       #tempPositionOfPostfix := #tempPositionOfPostfix + 1;
       #tempPositionOfPrePostfix := #tempPositionOfPrePostfix + 1;
       WHILE (#tempPrePostfix[#tempPositionOfPrePostfix + 1]) <= #LGCODE_MTH_PRSR_NUMBER_9 AND
         (#tempPrePostfix[#tempPositionOfPrePostfix + 1] >= #LGCODE_MTH_PRSR_NUMBER_0) AND
         (#tempPositionOfPrePostfix < #tempMaxPositionOfPrePostfix) DO
         #tempPostfixNotation[#tempPositionOfPostfix - 1] :=
         #tempPostfixNotation[#tempPositionOfPostfix - 1] + (#tempPrePostfix[#tempPositionOfPrePostfix + 1] - #LGCODE_MTH_PRSR_NUMBER_0)
         / #tempDenominatorDecimalNumbers;
         #tempPositionOfPrePostfix := #tempPositionOfPrePostfix + 1;
         #tempDenominatorDecimalNumbers := #tempDenominatorDecimalNumbers * 10;
       END_WHILE;
       #tempDenominatorDecimalNumbers := 10;
       //Falls negative Zahl
       IF #tempNextPostfixNumberIsNegative = TRUE THEN
         #tempPostfixNotation[#tempPositionOfPostfix - 1] := #tempPostfixNotation[#tempPositionOfPostfix - 1] * (-1);
         #tempNextPostfixNumberIsNegative := FALSE;
       END_IF;
       #tempPositionDecimalNumbers[#tempNumberOfDecimalNo] := #tempPositionOfPostfix - 1;
       #tempNumberOfDecimalNo := #tempNumberOfDecimalNo + 1;
     ELSIF
       //Zwei oder mehr Zahlen hintereinander erkennen und Zehner-, Hunderter-, Tausender- Stelle bilden
       (#tempPrePostfix[#tempPositionOfPrePostfix] <= #LGCODE_MTH_PRSR_NUMBER_9) AND
       (#tempPrePostfix[#tempPositionOfPrePostfix] >= #LGCODE_MTH_PRSR_NUMBER_0) AND
       (#tempPrePostfix[#tempPositionOfPrePostfix + 1] <= #LGCODE_MTH_PRSR_NUMBER_9) AND
       (#tempPrePostfix[#tempPositionOfPrePostfix + 1] >= #LGCODE_MTH_PRSR_NUMBER_0) AND
       (#tempPositionOfPrePostfix < #tempMaxPositionOfPrePostfix) AND
       (#tempPositionOfPrePostfix <> 0)
     THEN
       #tempPostfixNotation[#tempPositionOfPostfix] := (#tempPrePostfix[#tempPositionOfPrePostfix] - #LGCODE_MTH_PRSR_NUMBER_0);
       #tempPositionOfPostfix := #tempPositionOfPostfix + 1;
       WHILE (#tempPrePostfix[#tempPositionOfPrePostfix + 1] <= #LGCODE_MTH_PRSR_NUMBER_9) AND
         (#tempPrePostfix[#tempPositionOfPrePostfix + 1] >= #LGCODE_MTH_PRSR_NUMBER_0) AND
         (#tempPositionOfPrePostfix < #tempMaxPositionOfPrePostfix) DO
         #tempPostfixNotation[#tempPositionOfPostfix - 1] :=
         #tempPostfixNotation[#tempPositionOfPostfix - 1] * #LGCODE_MTH_PRSR_MULTIPLIER_FOR_MULTI_DIGIT_NO +
         (#tempPrePostfix[#tempPositionOfPrePostfix + 1] - #LGCODE_MTH_PRSR_NUMBER_0);
         #tempPositionOfPrePostfix := #tempPositionOfPrePostfix + 1;
       END_WHILE;
       #tempPositionMultiDigitNumbers[#tempNumberOfMultiDigitNo] := #tempPositionOfPostfix - 1;
       #tempNumberOfMultiDigitNo := #tempNumberOfMultiDigitNo + 1;
       //Falls mehrstellige Kommazahl
       IF #tempPrePostfix[#tempPositionOfPrePostfix + 1] = #LGCODE_MTH_PRSR_DECIMAL_POINT THEN
         #tempPositionOfPrePostfix := #tempPositionOfPrePostfix + 1;
         WHILE (#tempPrePostfix[#tempPositionOfPrePostfix + 1] <= #LGCODE_MTH_PRSR_NUMBER_9) AND
           (#tempPrePostfix[#tempPositionOfPrePostfix + 1] >= #LGCODE_MTH_PRSR_NUMBER_0) AND
           (#tempPositionOfPrePostfix < #tempMaxPositionOfPrePostfix) DO
           #tempPostfixNotation[#tempPositionOfPostfix - 1] := #tempPostfixNotation[#tempPositionOfPostfix - 1] +
           (#tempPrePostfix[#tempPositionOfPrePostfix + 1] - #LGCODE_MTH_PRSR_NUMBER_0) / #tempDenominatorDecimalNumbers;
           #tempPositionOfPrePostfix := #tempPositionOfPrePostfix + 1;
           #tempDenominatorDecimalNumbers := #tempDenominatorDecimalNumbers * 10;
         END_WHILE;
         #tempDenominatorDecimalNumbers := 10;
         #tempPositionDecimalNumbers[#tempNumberOfDecimalNo] := #tempPositionOfPostfix - 1;
         #tempNumberOfDecimalNo := #tempNumberOfDecimalNo + 1;
       END_IF;
       //Falls negative Zahl
       IF #tempNextPostfixNumberIsNegative = TRUE THEN
         #tempPostfixNotation[#tempPositionOfPostfix - 1] := #tempPostfixNotation[#tempPositionOfPostfix - 1] * (-1);
         #tempNextPostfixNumberIsNegative := FALSE;
       END_IF;
     ELSIF
       //Zahlen in Postfix-Notation schreiben
       (#tempPrePostfix[#tempPositionOfPrePostfix] <= #LGCODE_MTH_PRSR_NUMBER_9) AND (#tempPrePostfix[#tempPositionOfPrePostfix] >= #LGCODE_MTH_PRSR_NUMBER_0)
     THEN
       #tempPostfixNotation[#tempPositionOfPostfix] := (#tempPrePostfix[#tempPositionOfPrePostfix] - #LGCODE_MTH_PRSR_NUMBER_0);
       #tempPositionOfPostfix := #tempPositionOfPostfix + 1;
       //Falls negative Zahl
       IF #tempNextPostfixNumberIsNegative = TRUE THEN
         #tempPostfixNotation[#tempPositionOfPostfix - 1] := #tempPostfixNotation[#tempPositionOfPostfix - 1] * (-1);
         #tempNextPostfixNumberIsNegative := FALSE;
       END_IF;
     ELSIF
       //negative Zahlen erkennen
       ((#tempPrePostfix[#tempPositionOfPrePostfix] = #LGCODE_MTH_PRSR_MINUS) AND

       ((#tempPrePostfix[#tempPositionOfPrePostfix + 1] >= #LGCODE_MTH_PRSR_NUMBER_0) AND
       (#tempPrePostfix[#tempPositionOfPrePostfix + 1] <= #LGCODE_MTH_PRSR_NUMBER_9)) AND

       ((#tempPrePostfix[#tempPositionOfPrePostfix - 1] = #LGCODE_MTH_PRSR_MINUS) OR
       (#tempPrePostfix[#tempPositionOfPrePostfix - 1] = #LGCODE_MTH_PRSR_TIMES) OR
       (#tempPrePostfix[#tempPositionOfPrePostfix - 1] = #LGCODE_MTH_PRSR_PLUS) OR
       (#tempPrePostfix[#tempPositionOfPrePostfix - 1] = #LGCODE_MTH_PRSR_MINUS) OR
       (#tempPrePostfix[#tempPositionOfPrePostfix - 1] = #LGCODE_MTH_PRSR_DIVIDE) OR
       (#tempPrePostfix[#tempPositionOfPrePostfix - 1] = #LGCODE_MTH_PRSR_OPEN_BRACKET) OR
       (#tempPrePostfix[#tempPositionOfPrePostfix - 1] = #LGCODE_MTH_PRSR_LOGICAL_OR) OR
       (#tempPrePostfix[#tempPositionOfPrePostfix - 1] = #LGCODE_MTH_PRSR_LOGICAL_AND) OR
       (#tempPrePostfix[#tempPositionOfPrePostfix - 1] = #LGCODE_MTH_PRSR_LOGICAL_GREATER) OR
       (#tempPrePostfix[#tempPositionOfPrePostfix - 1] = #LGCODE_MTH_PRSR_LOGICAL_LESS) OR
       (#tempPrePostfix[#tempPositionOfPrePostfix - 1] = #LGCODE_MTH_PRSR_LOGICAL_EQUAL) OR
       (#tempPrePostfix[#tempPositionOfPrePostfix - 1] = #LGCODE_MTH_PRSR_LOGICAL_GREATER_EQUAL) OR
       (#tempPrePostfix[#tempPositionOfPrePostfix - 1] = #LGCODE_MTH_PRSR_LOGICAL_LESS_EQUAL) OR
       (#tempPrePostfix[#tempPositionOfPrePostfix - 1] = #LGCODE_MTH_PRSR_LOGICAL_NOT_EQUAL) OR
       (#tempPrePostfix[#tempPositionOfPrePostfix - 1] = #LGCODE_MTH_PRSR_LOGICAL_NOT) OR
       (#tempPrePostfix[#tempPositionOfPrePostfix - 1] = #LGCODE_MTH_PRSR_TO_THE_POWER_OF) OR
       (#tempPositionOfPrePostfix = 1)))
     THEN
       #tempNextPostfixNumberIsNegative := TRUE;
     ELSIF
       //negative Klammerausdrücke erkennen
       (#tempPrePostfix[#tempPositionOfPrePostfix] = #LGCODE_MTH_PRSR_MINUS) AND

       (#tempPrePostfix[#tempPositionOfPrePostfix + 1] = #LGCODE_MTH_PRSR_OPEN_BRACKET) AND

       ((#tempPrePostfix[#tempPositionOfPrePostfix - 1] = #LGCODE_MTH_PRSR_TIMES) OR
       (#tempPrePostfix[#tempPositionOfPrePostfix - 1] = #LGCODE_MTH_PRSR_PLUS) OR
       (#tempPrePostfix[#tempPositionOfPrePostfix - 1] = #LGCODE_MTH_PRSR_MINUS) OR
       (#tempPrePostfix[#tempPositionOfPrePostfix - 1] = #LGCODE_MTH_PRSR_DIVIDE) OR
       (#tempPrePostfix[#tempPositionOfPrePostfix - 1] = #LGCODE_MTH_PRSR_OPEN_BRACKET) OR
       (#tempPrePostfix[#tempPositionOfPrePostfix - 1] = #LGCODE_MTH_PRSR_CHAR_N) OR
       (#tempPrePostfix[#tempPositionOfPrePostfix - 1] = #LGCODE_MTH_PRSR_CHAR_S) OR
       (#tempPrePostfix[#tempPositionOfPrePostfix - 1] = #LGCODE_MTH_PRSR_CHAR_R) OR
       (#tempPrePostfix[#tempPositionOfPrePostfix - 1] = #LGCODE_MTH_PRSR_CHAR_T) OR
       (#tempPrePostfix[#tempPositionOfPrePostfix - 1] = #LGCODE_MTH_PRSR_LOGICAL_OR) OR
       (#tempPrePostfix[#tempPositionOfPrePostfix - 1] = #LGCODE_MTH_PRSR_LOGICAL_AND) OR
       (#tempPrePostfix[#tempPositionOfPrePostfix - 1] = #LGCODE_MTH_PRSR_LOGICAL_GREATER) OR
       (#tempPrePostfix[#tempPositionOfPrePostfix - 1] = #LGCODE_MTH_PRSR_LOGICAL_LESS) OR
       (#tempPrePostfix[#tempPositionOfPrePostfix - 1] = #LGCODE_MTH_PRSR_LOGICAL_EQUAL) OR
       (#tempPrePostfix[#tempPositionOfPrePostfix - 1] = #LGCODE_MTH_PRSR_LOGICAL_GREATER_EQUAL) OR
       (#tempPrePostfix[#tempPositionOfPrePostfix - 1] = #LGCODE_MTH_PRSR_LOGICAL_LESS_EQUAL) OR
       (#tempPrePostfix[#tempPositionOfPrePostfix - 1] = #LGCODE_MTH_PRSR_LOGICAL_NOT_EQUAL) OR
       (#tempPrePostfix[#tempPositionOfPrePostfix - 1] = #LGCODE_MTH_PRSR_LOGICAL_NOT) OR
       (#tempPrePostfix[#tempPositionOfPrePostfix - 1] = #LGCODE_MTH_PRSR_TO_THE_POWER_OF) OR
       (#tempPositionOfPrePostfix = 1))
     THEN
       #tempPositionOfNegBrackets[#tempNumberOfNegBrackets] := #tempPositionOfOperatorStack;
       #tempNumberOfNegBrackets := #tempNumberOfNegBrackets + 1;
     ELSIF
       //negative mathematische Funktion erkennen
       (#tempPrePostfix[#tempPositionOfPrePostfix] = #LGCODE_MTH_PRSR_MINUS) AND

       ((#tempPrePostfix[#tempPositionOfPrePostfix + 1] = #LGCODE_MTH_PRSR_CHAR_C) OR
       (#tempPrePostfix[#tempPositionOfPrePostfix + 1] = #LGCODE_MTH_PRSR_CHAR_S)) AND

       ((#tempPrePostfix[#tempPositionOfPrePostfix - 1] = #LGCODE_MTH_PRSR_TIMES) OR
       (#tempPrePostfix[#tempPositionOfPrePostfix - 1] = #LGCODE_MTH_PRSR_PLUS) OR
       (#tempPrePostfix[#tempPositionOfPrePostfix - 1] = #LGCODE_MTH_PRSR_MINUS) OR
       (#tempPrePostfix[#tempPositionOfPrePostfix - 1] = #LGCODE_MTH_PRSR_DIVIDE) OR
       (#tempPrePostfix[#tempPositionOfPrePostfix - 1] = #LGCODE_MTH_PRSR_OPEN_BRACKET) OR
       (#tempPrePostfix[#tempPositionOfPrePostfix - 1] = #LGCODE_MTH_PRSR_LOGICAL_OR) OR
       (#tempPrePostfix[#tempPositionOfPrePostfix - 1] = #LGCODE_MTH_PRSR_LOGICAL_AND) OR
       (#tempPrePostfix[#tempPositionOfPrePostfix - 1] = #LGCODE_MTH_PRSR_LOGICAL_GREATER) OR
       (#tempPrePostfix[#tempPositionOfPrePostfix - 1] = #LGCODE_MTH_PRSR_LOGICAL_LESS) OR
       (#tempPrePostfix[#tempPositionOfPrePostfix - 1] = #LGCODE_MTH_PRSR_LOGICAL_EQUAL) OR
       (#tempPrePostfix[#tempPositionOfPrePostfix - 1] = #LGCODE_MTH_PRSR_LOGICAL_GREATER_EQUAL) OR
       (#tempPrePostfix[#tempPositionOfPrePostfix - 1] = #LGCODE_MTH_PRSR_LOGICAL_LESS_EQUAL) OR
       (#tempPrePostfix[#tempPositionOfPrePostfix - 1] = #LGCODE_MTH_PRSR_LOGICAL_NOT_EQUAL) OR
       (#tempPrePostfix[#tempPositionOfPrePostfix - 1] = #LGCODE_MTH_PRSR_LOGICAL_NOT) OR
       (#tempPrePostfix[#tempPositionOfPrePostfix - 1] = #LGCODE_MTH_PRSR_TO_THE_POWER_OF) OR
       (#tempPositionOfPrePostfix = 1))
     THEN
       #tempPositionOfNegFunctions[#tempNumberOfNegFunctions] := #tempPositionOfOperatorStack;
       #tempNumberOfNegFunctions := #tempNumberOfNegFunctions + 1;
     ELSIF
       //Zeichen je nach Bedingungen in Zeichenspeicher oder in Postfix-Notation schreiben
       //Zeichenspeicher leer, Zeichen in Zeichenspeicher schreiben
       (((#tempPrePostfix[#tempPositionOfPrePostfix] = #LGCODE_MTH_PRSR_LOGICAL_OR) OR
       (#tempPrePostfix[#tempPositionOfPrePostfix] = #LGCODE_MTH_PRSR_LOGICAL_AND) OR
       (#tempPrePostfix[#tempPositionOfPrePostfix] = #LGCODE_MTH_PRSR_LOGICAL_GREATER) OR
       (#tempPrePostfix[#tempPositionOfPrePostfix] = #LGCODE_MTH_PRSR_LOGICAL_LESS) OR
       (#tempPrePostfix[#tempPositionOfPrePostfix] = #LGCODE_MTH_PRSR_LOGICAL_EQUAL) OR
       (#tempPrePostfix[#tempPositionOfPrePostfix] = #LGCODE_MTH_PRSR_LOGICAL_GREATER_EQUAL) OR
       (#tempPrePostfix[#tempPositionOfPrePostfix] = #LGCODE_MTH_PRSR_LOGICAL_LESS_EQUAL) OR
       (#tempPrePostfix[#tempPositionOfPrePostfix] = #LGCODE_MTH_PRSR_LOGICAL_NOT_EQUAL) OR
       (#tempPrePostfix[#tempPositionOfPrePostfix] = #LGCODE_MTH_PRSR_LOGICAL_NOT) OR
       (#tempPrePostfix[#tempPositionOfPrePostfix] = #LGCODE_MTH_PRSR_TIMES) OR
       (#tempPrePostfix[#tempPositionOfPrePostfix] = #LGCODE_MTH_PRSR_DIVIDE) OR
       (#tempPrePostfix[#tempPositionOfPrePostfix] = #LGCODE_MTH_PRSR_PLUS) OR
       (#tempPrePostfix[#tempPositionOfPrePostfix] = #LGCODE_MTH_PRSR_MINUS)) AND
       (#tempPositionOfOperatorStack = 1))
     THEN
       #tempStackForOperators[#tempPositionOfOperatorStack] := #tempPrePostfix[#tempPositionOfPrePostfix];
       #tempPositionOfOperatorStack := #tempPositionOfOperatorStack + 1;
     ELSIF
       //letztes Zeichen boolesch und nächstes mathematisch
       //Zeichen in Zeichenspeicher speichern
       ((#tempStackForOperators[#tempPositionOfOperatorStack - 1] = #LGCODE_MTH_PRSR_LOGICAL_GREATER) OR
       (#tempStackForOperators[#tempPositionOfOperatorStack - 1] = #LGCODE_MTH_PRSR_LOGICAL_LESS) OR
       (#tempStackForOperators[#tempPositionOfOperatorStack - 1] = #LGCODE_MTH_PRSR_LOGICAL_GREATER_EQUAL) OR
       (#tempStackForOperators[#tempPositionOfOperatorStack - 1] = #LGCODE_MTH_PRSR_LOGICAL_LESS_EQUAL) OR
       (#tempStackForOperators[#tempPositionOfOperatorStack - 1] = #LGCODE_MTH_PRSR_LOGICAL_EQUAL) OR
       (#tempStackForOperators[#tempPositionOfOperatorStack - 1] = #LGCODE_MTH_PRSR_LOGICAL_NOT_EQUAL) OR
       (#tempStackForOperators[#tempPositionOfOperatorStack - 1] = #LGCODE_MTH_PRSR_LOGICAL_AND) OR
       (#tempStackForOperators[#tempPositionOfOperatorStack - 1] = #LGCODE_MTH_PRSR_LOGICAL_OR))
       AND
       ((#tempPrePostfix[#tempPositionOfPrePostfix] = #LGCODE_MTH_PRSR_PLUS) OR
       (#tempPrePostfix[#tempPositionOfPrePostfix] = #LGCODE_MTH_PRSR_MINUS) OR
       (#tempPrePostfix[#tempPositionOfPrePostfix] = #LGCODE_MTH_PRSR_TIMES) OR
       (#tempPrePostfix[#tempPositionOfPrePostfix] = #LGCODE_MTH_PRSR_DIVIDE) OR
       (#tempPrePostfix[#tempPositionOfPrePostfix] = #LGCODE_MTH_PRSR_OPEN_BRACKET))
     THEN
       #tempStackForOperators[#tempPositionOfOperatorStack] := #tempPrePostfix[#tempPositionOfPrePostfix];
       #tempPositionOfOperatorStack := #tempPositionOfOperatorStack + 1;
     ELSIF
       //letztes Zeichen mathematisch und nächstes boolesch
       //dann alle mathematischen Zeichen erst aus Zeichenspeicher holen
       ((#tempStackForOperators[#tempPositionOfOperatorStack - 1] = #LGCODE_MTH_PRSR_TIMES) OR
       (#tempStackForOperators[#tempPositionOfOperatorStack - 1] = #LGCODE_MTH_PRSR_DIVIDE) OR
       (#tempStackForOperators[#tempPositionOfOperatorStack - 1] = #LGCODE_MTH_PRSR_MINUS) OR
       (#tempStackForOperators[#tempPositionOfOperatorStack - 1] = #LGCODE_MTH_PRSR_PLUS) OR
       (#tempStackForOperators[#tempPositionOfOperatorStack - 1] = #LGCODE_MTH_PRSR_SINUS) OR
       (#tempStackForOperators[#tempPositionOfOperatorStack - 1] = #LGCODE_MTH_PRSR_COSINUS) OR
       (#tempStackForOperators[#tempPositionOfOperatorStack - 1] = #LGCODE_MTH_PRSR_SQUARE) OR
       (#tempStackForOperators[#tempPositionOfOperatorStack - 1] = #LGCODE_MTH_PRSR_SQUAREROOT))
       AND
       ((#tempPrePostfix[#tempPositionOfPrePostfix] = #LGCODE_MTH_PRSR_LOGICAL_GREATER_EQUAL) OR
       (#tempPrePostfix[#tempPositionOfPrePostfix] = #LGCODE_MTH_PRSR_LOGICAL_LESS_EQUAL) OR
       (#tempPrePostfix[#tempPositionOfPrePostfix] = #LGCODE_MTH_PRSR_LOGICAL_EQUAL) OR
       (#tempPrePostfix[#tempPositionOfPrePostfix] = #LGCODE_MTH_PRSR_LOGICAL_NOT_EQUAL) OR
       (#tempPrePostfix[#tempPositionOfPrePostfix] = #LGCODE_MTH_PRSR_LOGICAL_GREATER) OR
       (#tempPrePostfix[#tempPositionOfPrePostfix] = #LGCODE_MTH_PRSR_LOGICAL_LESS) OR
       (#tempPrePostfix[#tempPositionOfPrePostfix] = #LGCODE_MTH_PRSR_LOGICAL_AND) OR
       (#tempPrePostfix[#tempPositionOfPrePostfix] = #LGCODE_MTH_PRSR_LOGICAL_OR))
     THEN
       #tempPostfixNotation[#tempPositionOfPostfix] := #tempStackForOperators[#tempPositionOfOperatorStack - 1];
       #tempPositionOfPostfix := #tempPositionOfPostfix + 1;
       #tempPositionOfOperatorStack := #tempPositionOfOperatorStack - 1;
       IF (#tempStackForOperators[#tempPositionOfOperatorStack - 1] = #LGCODE_MTH_PRSR_PLUS) OR
         (#tempStackForOperators[#tempPositionOfOperatorStack - 1] = #LGCODE_MTH_PRSR_MINUS) OR
         (#tempStackForOperators[#tempPositionOfOperatorStack - 1] = #LGCODE_MTH_PRSR_TIMES) OR
         (#tempStackForOperators[#tempPositionOfOperatorStack - 1] = #LGCODE_MTH_PRSR_DIVIDE)
       THEN
         #tempPostfixNotation[#tempPositionOfPostfix] := #tempStackForOperators[#tempPositionOfOperatorStack - 1];
         #tempPositionOfPostfix := #tempPositionOfPostfix + 1;
         #tempPositionOfOperatorStack := #tempPositionOfOperatorStack - 1;
       END_IF;
       #tempStackForOperators[#tempPositionOfOperatorStack] := #tempPrePostfix[#tempPositionOfPrePostfix];
       #tempPositionOfOperatorStack := #tempPositionOfOperatorStack + 1;
     ELSIF
       //letztes Zeichen >/ >= / <=/ =/<> oder < Nächstes & oder | dann Zeichen erst aus Zeichenspeicher holen
       ((#tempStackForOperators[#tempPositionOfOperatorStack - 1] = #LGCODE_MTH_PRSR_LOGICAL_GREATER) OR
       (#tempStackForOperators[#tempPositionOfOperatorStack - 1] = #LGCODE_MTH_PRSR_LOGICAL_LESS) OR
       (#tempStackForOperators[#tempPositionOfOperatorStack - 1] = #LGCODE_MTH_PRSR_LOGICAL_GREATER_EQUAL) OR
       (#tempStackForOperators[#tempPositionOfOperatorStack - 1] = #LGCODE_MTH_PRSR_LOGICAL_LESS_EQUAL) OR
       (#tempStackForOperators[#tempPositionOfOperatorStack - 1] = #LGCODE_MTH_PRSR_LOGICAL_EQUAL) OR
       (#tempStackForOperators[#tempPositionOfOperatorStack - 1] = #LGCODE_MTH_PRSR_LOGICAL_NOT_EQUAL))
       AND
       ((#tempPrePostfix[#tempPositionOfPrePostfix] = #LGCODE_MTH_PRSR_LOGICAL_AND) OR
       (#tempPrePostfix[#tempPositionOfPrePostfix] = #LGCODE_MTH_PRSR_LOGICAL_OR))
     THEN
       #tempPostfixNotation[#tempPositionOfPostfix] := #tempStackForOperators[#tempPositionOfOperatorStack - 1];
       #tempPositionOfPostfix := #tempPositionOfPostfix + 1;
       #tempPositionOfOperatorStack := #tempPositionOfOperatorStack - 1;
       IF    //Falls nächstes Zeichen im Zeichenspeicher noch ein AND oder AND
         ((#tempStackForOperators[#tempPositionOfOperatorStack - 1] = #LGCODE_MTH_PRSR_LOGICAL_AND) OR
         (#tempStackForOperators[#tempPositionOfOperatorStack - 1] = #LGCODE_MTH_PRSR_LOGICAL_OR))
       THEN
         #tempPostfixNotation[#tempPositionOfPostfix] := #tempStackForOperators[#tempPositionOfOperatorStack - 1];
         #tempPositionOfPostfix := #tempPositionOfPostfix + 1;
         #tempPositionOfOperatorStack := #tempPositionOfOperatorStack - 1;
       END_IF;
       #tempStackForOperators[#tempPositionOfOperatorStack] := #tempPrePostfix[#tempPositionOfPrePostfix];
       #tempPositionOfOperatorStack := #tempPositionOfOperatorStack + 1;
     ELSIF
       //letztes Zeichen >/ < / >=/<= /<> /=  oder <  und Nächstes ein >/ >= / <=/ <>/ = oder < dann erst Zeichen aus Zeichenspeicher holen
       //und dann erst kommendes Zeichen in Stack schreiben
       ((#tempStackForOperators[#tempPositionOfOperatorStack - 1] = #LGCODE_MTH_PRSR_LOGICAL_GREATER) OR
       (#tempStackForOperators[#tempPositionOfOperatorStack - 1] = #LGCODE_MTH_PRSR_LOGICAL_LESS) OR
       (#tempStackForOperators[#tempPositionOfOperatorStack - 1] = #LGCODE_MTH_PRSR_LOGICAL_GREATER_EQUAL) OR
       (#tempStackForOperators[#tempPositionOfOperatorStack - 1] = #LGCODE_MTH_PRSR_LOGICAL_LESS_EQUAL) OR
       (#tempStackForOperators[#tempPositionOfOperatorStack - 1] = #LGCODE_MTH_PRSR_LOGICAL_NOT_EQUAL) OR
       (#tempStackForOperators[#tempPositionOfOperatorStack - 1] = #LGCODE_MTH_PRSR_LOGICAL_EQUAL))
       AND
       ((#tempPrePostfix[#tempPositionOfPrePostfix] = #LGCODE_MTH_PRSR_LOGICAL_GREATER) OR
       (#tempPrePostfix[#tempPositionOfPrePostfix] = #LGCODE_MTH_PRSR_LOGICAL_LESS) OR
       (#tempPrePostfix[#tempPositionOfPrePostfix] = #LGCODE_MTH_PRSR_LOGICAL_GREATER_EQUAL) OR
       (#tempPrePostfix[#tempPositionOfPrePostfix] = #LGCODE_MTH_PRSR_LOGICAL_LESS_EQUAL) OR
       (#tempPrePostfix[#tempPositionOfPrePostfix] = #LGCODE_MTH_PRSR_LOGICAL_NOT_EQUAL) OR
       (#tempPrePostfix[#tempPositionOfPrePostfix] = #LGCODE_MTH_PRSR_LOGICAL_EQUAL))
     THEN
       #tempPostfixNotation[#tempPositionOfPostfix] := #tempStackForOperators[#tempPositionOfOperatorStack - 1];
       #tempPositionOfPostfix := #tempPositionOfPostfix + 1;
       #tempPositionOfOperatorStack := #tempPositionOfOperatorStack - 1;
       #tempStackForOperators[#tempPositionOfOperatorStack] := #tempPrePostfix[#tempPositionOfPrePostfix];
       #tempPositionOfOperatorStack := #tempPositionOfOperatorStack + 1;
     ELSIF
       //letztes Zeichen & oder | und Nächstes > /< />= / <= /<> /=   oder < dann Zeichen in Zeichenspeicher schreiben
       ((#tempStackForOperators[#tempPositionOfOperatorStack - 1] = #LGCODE_MTH_PRSR_LOGICAL_AND) OR
       (#tempStackForOperators[#tempPositionOfOperatorStack - 1] = #LGCODE_MTH_PRSR_LOGICAL_OR))
       AND
       ((#tempPrePostfix[#tempPositionOfPrePostfix] = #LGCODE_MTH_PRSR_LOGICAL_GREATER) OR
       (#tempPrePostfix[#tempPositionOfPrePostfix] = #LGCODE_MTH_PRSR_LOGICAL_LESS) OR
       (#tempPrePostfix[#tempPositionOfPrePostfix] = #LGCODE_MTH_PRSR_LOGICAL_GREATER_EQUAL) OR
       (#tempPrePostfix[#tempPositionOfPrePostfix] = #LGCODE_MTH_PRSR_LOGICAL_LESS_EQUAL) OR
       (#tempPrePostfix[#tempPositionOfPrePostfix] = #LGCODE_MTH_PRSR_LOGICAL_NOT_EQUAL) OR
       (#tempPrePostfix[#tempPositionOfPrePostfix] = #LGCODE_MTH_PRSR_LOGICAL_EQUAL))
     THEN
       #tempStackForOperators[#tempPositionOfOperatorStack] := #tempPrePostfix[#tempPositionOfPrePostfix];
       #tempPositionOfOperatorStack := #tempPositionOfOperatorStack + 1;
     ELSIF
       //letztes Zeichen  & oder | und Nächstes & oder | dann Zeichen erst aus Zeichenspeicher holen
       ((#tempStackForOperators[#tempPositionOfOperatorStack - 1] = #LGCODE_MTH_PRSR_LOGICAL_AND) OR
       (#tempStackForOperators[#tempPositionOfOperatorStack - 1] = #LGCODE_MTH_PRSR_LOGICAL_OR))
       AND
       ((#tempPrePostfix[#tempPositionOfPrePostfix] = #LGCODE_MTH_PRSR_LOGICAL_AND) OR
       (#tempPrePostfix[#tempPositionOfPrePostfix] = #LGCODE_MTH_PRSR_LOGICAL_OR))
     THEN
       #tempPostfixNotation[#tempPositionOfPostfix] := #tempStackForOperators[#tempPositionOfOperatorStack - 1];
       #tempPositionOfPostfix := #tempPositionOfPostfix + 1;
       #tempPositionOfOperatorStack := #tempPositionOfOperatorStack - 1;
       #tempStackForOperators[#tempPositionOfOperatorStack] := #tempPrePostfix[#tempPositionOfPrePostfix];
       #tempPositionOfOperatorStack := #tempPositionOfOperatorStack + 1;

     ELSIF
       //! immer in Zeichenspeicher schreiben
       (#tempPrePostfix[#tempPositionOfPrePostfix] = #LGCODE_MTH_PRSR_LOGICAL_NOT)
     THEN
       #tempStackForOperators[#tempPositionOfOperatorStack] := #tempPrePostfix[#tempPositionOfPrePostfix];
       #tempPositionOfOperatorStack := #tempPositionOfOperatorStack + 1;
     ELSIF
       //bei kommenden Zeichen, ! aus Zeichenspeicher holen
       (#tempStackForOperators[#tempPositionOfOperatorStack - 1] = #LGCODE_MTH_PRSR_LOGICAL_NOT)
       AND
       ((#tempPrePostfix[#tempPositionOfPrePostfix] = #LGCODE_MTH_PRSR_LOGICAL_GREATER) OR
       (#tempPrePostfix[#tempPositionOfPrePostfix] = #LGCODE_MTH_PRSR_LOGICAL_LESS) OR
       (#tempPrePostfix[#tempPositionOfPrePostfix] = #LGCODE_MTH_PRSR_LOGICAL_GREATER_EQUAL) OR
       (#tempPrePostfix[#tempPositionOfPrePostfix] = #LGCODE_MTH_PRSR_LOGICAL_LESS_EQUAL) OR
       (#tempPrePostfix[#tempPositionOfPrePostfix] = #LGCODE_MTH_PRSR_LOGICAL_NOT_EQUAL) OR
       (#tempPrePostfix[#tempPositionOfPrePostfix] = #LGCODE_MTH_PRSR_LOGICAL_EQUAL) OR
       (#tempPrePostfix[#tempPositionOfPrePostfix] = #LGCODE_MTH_PRSR_LOGICAL_AND) OR
       (#tempPrePostfix[#tempPositionOfPrePostfix] = #LGCODE_MTH_PRSR_LOGICAL_OR) OR
       (#tempPrePostfix[#tempPositionOfPrePostfix] = #LGCODE_MTH_PRSR_TO_THE_POWER_OF) OR
       (#tempPrePostfix[#tempPositionOfPrePostfix] = #LGCODE_MTH_PRSR_PLUS) OR
       (#tempPrePostfix[#tempPositionOfPrePostfix] = #LGCODE_MTH_PRSR_MINUS) OR
       (#tempPrePostfix[#tempPositionOfPrePostfix] = #LGCODE_MTH_PRSR_TIMES) OR
       (#tempPrePostfix[#tempPositionOfPrePostfix] = #LGCODE_MTH_PRSR_DIVIDE) OR
       (#tempPrePostfix[#tempPositionOfPrePostfix] = #LGCODE_MTH_PRSR_SINUS) OR
       (#tempPrePostfix[#tempPositionOfPrePostfix] = #LGCODE_MTH_PRSR_COSINUS) OR
       (#tempPrePostfix[#tempPositionOfPrePostfix] = #LGCODE_MTH_PRSR_SQUARE) OR
       (#tempPrePostfix[#tempPositionOfPrePostfix] = #LGCODE_MTH_PRSR_SQUAREROOT))
     THEN
       #tempPostfixNotation[#tempPositionOfPostfix] := #tempStackForOperators[#tempPositionOfOperatorStack - 1];
       #tempPositionOfPostfix := #tempPositionOfPostfix + 1;
       #tempPositionOfOperatorStack := #tempPositionOfOperatorStack - 1;
       //damit ausräumendes Zeichen im nächsten Durchgang korrekt verarbeitet wird
       #tempPositionOfPrePostfix := #tempPositionOfPrePostfix - 1;
     ELSIF
       //^ (Exponential-Operator) bei nächstem Zeichen aus Zeichenspeicher holen
       ((#tempStackForOperators[#tempPositionOfOperatorStack - 1] = #LGCODE_MTH_PRSR_TO_THE_POWER_OF)
       AND
       ((#tempPrePostfix[#tempPositionOfPrePostfix] = #LGCODE_MTH_PRSR_LOGICAL_GREATER) OR
       (#tempPrePostfix[#tempPositionOfPrePostfix] = #LGCODE_MTH_PRSR_LOGICAL_LESS) OR
       (#tempPrePostfix[#tempPositionOfPrePostfix] = #LGCODE_MTH_PRSR_LOGICAL_GREATER_EQUAL) OR
       (#tempPrePostfix[#tempPositionOfPrePostfix] = #LGCODE_MTH_PRSR_LOGICAL_LESS_EQUAL) OR
       (#tempPrePostfix[#tempPositionOfPrePostfix] = #LGCODE_MTH_PRSR_LOGICAL_NOT_EQUAL) OR
       (#tempPrePostfix[#tempPositionOfPrePostfix] = #LGCODE_MTH_PRSR_LOGICAL_EQUAL) OR
       (#tempPrePostfix[#tempPositionOfPrePostfix] = #LGCODE_MTH_PRSR_LOGICAL_AND) OR
       (#tempPrePostfix[#tempPositionOfPrePostfix] = #LGCODE_MTH_PRSR_LOGICAL_OR) OR
       (#tempPrePostfix[#tempPositionOfPrePostfix] = #LGCODE_MTH_PRSR_TO_THE_POWER_OF) OR
       (#tempPrePostfix[#tempPositionOfPrePostfix] = #LGCODE_MTH_PRSR_PLUS) OR
       (#tempPrePostfix[#tempPositionOfPrePostfix] = #LGCODE_MTH_PRSR_MINUS) OR
       (#tempPrePostfix[#tempPositionOfPrePostfix] = #LGCODE_MTH_PRSR_TIMES) OR
       (#tempPrePostfix[#tempPositionOfPrePostfix] = #LGCODE_MTH_PRSR_DIVIDE)))
     THEN
       #tempPostfixNotation[#tempPositionOfPostfix] := #tempStackForOperators[#tempPositionOfOperatorStack - 1];
       #tempPositionOfPostfix := #tempPositionOfPostfix + 1;
       #tempPositionOfOperatorStack := #tempPositionOfOperatorStack - 1;
       //damit ausräumendes Zeichen im nächsten Durchgang korrekt verarbeitet wird
       #tempPositionOfPrePostfix := #tempPositionOfPrePostfix - 1;
     ELSIF
       //^ (Exponential-Operator) in Zeichenspeicher schreiben,
       //außer oberstes Zeichen ist Funktion oder NOT, ist weiter oben realisiert
       (#tempPrePostfix[#tempPositionOfPrePostfix] = #LGCODE_MTH_PRSR_TO_THE_POWER_OF)
     THEN
       #tempStackForOperators[#tempPositionOfOperatorStack] := #tempPrePostfix[#tempPositionOfPrePostfix];
       #tempPositionOfOperatorStack := #tempPositionOfOperatorStack + 1;
     ELSIF
       //letztes Zeichen * oder / Nächstes + oder - dann erst Zeichen aus Zeichenspeicher holen
       ((#tempStackForOperators[#tempPositionOfOperatorStack - 1] = #LGCODE_MTH_PRSR_TIMES) OR
       (#tempStackForOperators[#tempPositionOfOperatorStack - 1] = #LGCODE_MTH_PRSR_DIVIDE)) AND
       ((#tempPrePostfix[#tempPositionOfPrePostfix] = #LGCODE_MTH_PRSR_PLUS) OR
       (#tempPrePostfix[#tempPositionOfPrePostfix] = #LGCODE_MTH_PRSR_MINUS))
     THEN
       #tempPostfixNotation[#tempPositionOfPostfix] := #tempStackForOperators[#tempPositionOfOperatorStack - 1];
       #tempPositionOfPostfix := #tempPositionOfPostfix + 1;
       #tempPositionOfOperatorStack := #tempPositionOfOperatorStack - 1;
       IF    //Falls nächstes Zeichen im Zeichenspeicher noch ein + oder -
         ((#tempStackForOperators[#tempPositionOfOperatorStack - 1] = #LGCODE_MTH_PRSR_PLUS) OR
         (#tempStackForOperators[#tempPositionOfOperatorStack - 1] = #LGCODE_MTH_PRSR_MINUS))
       THEN
         #tempPostfixNotation[#tempPositionOfPostfix] := #tempStackForOperators[#tempPositionOfOperatorStack - 1];
         #tempPositionOfPostfix := #tempPositionOfPostfix + 1;
         #tempPositionOfOperatorStack := #tempPositionOfOperatorStack - 1;
       END_IF;
       #tempStackForOperators[#tempPositionOfOperatorStack] := #tempPrePostfix[#tempPositionOfPrePostfix];
       #tempPositionOfOperatorStack := #tempPositionOfOperatorStack + 1;
     ELSIF
       //letztes Zeichen  * oder / Nächstes ein * oder / dann erst Zeichen aus Zeichenspeicher holen
       //und dann erst kommendes Zeichen in Stack schreiben
       ((#tempStackForOperators[#tempPositionOfOperatorStack - 1] = #LGCODE_MTH_PRSR_TIMES) OR
       (#tempStackForOperators[#tempPositionOfOperatorStack - 1] = #LGCODE_MTH_PRSR_DIVIDE)) AND
       ((#tempPrePostfix[#tempPositionOfPrePostfix] = #LGCODE_MTH_PRSR_TIMES) OR
       (#tempPrePostfix[#tempPositionOfPrePostfix] = #LGCODE_MTH_PRSR_DIVIDE))
     THEN
       #tempPostfixNotation[#tempPositionOfPostfix] := #tempStackForOperators[#tempPositionOfOperatorStack - 1];
       #tempPositionOfPostfix := #tempPositionOfPostfix + 1;
       #tempPositionOfOperatorStack := #tempPositionOfOperatorStack - 1;
       #tempStackForOperators[#tempPositionOfOperatorStack] := #tempPrePostfix[#tempPositionOfPrePostfix];
       #tempPositionOfOperatorStack := #tempPositionOfOperatorStack + 1;
     ELSIF
       //letztes Zeichen ein + oder - und Nächstes * oder / dann Zeichen in Zeichenspeicher schreiben
       ((#tempStackForOperators[#tempPositionOfOperatorStack - 1] = #LGCODE_MTH_PRSR_PLUS) OR
       (#tempStackForOperators[#tempPositionOfOperatorStack - 1] = #LGCODE_MTH_PRSR_MINUS)) AND
       ((#tempPrePostfix[#tempPositionOfPrePostfix] = #LGCODE_MTH_PRSR_TIMES) OR
       (#tempPrePostfix[#tempPositionOfPrePostfix] = #LGCODE_MTH_PRSR_DIVIDE))
     THEN
       #tempStackForOperators[#tempPositionOfOperatorStack] := #tempPrePostfix[#tempPositionOfPrePostfix];
       #tempPositionOfOperatorStack := #tempPositionOfOperatorStack + 1;
     ELSIF
       //letztes Zeichen  + oder - und Nächstes + oder - dann Zeichen erst aus Zeichenspeicher holen
       ((#tempStackForOperators[#tempPositionOfOperatorStack - 1] = #LGCODE_MTH_PRSR_PLUS) OR
       (#tempStackForOperators[#tempPositionOfOperatorStack - 1] = #LGCODE_MTH_PRSR_MINUS)) AND
       ((#tempPrePostfix[#tempPositionOfPrePostfix] = #LGCODE_MTH_PRSR_PLUS) OR
       (#tempPrePostfix[#tempPositionOfPrePostfix] = #LGCODE_MTH_PRSR_MINUS))
     THEN
       #tempPostfixNotation[#tempPositionOfPostfix] := #tempStackForOperators[#tempPositionOfOperatorStack - 1];
       #tempPositionOfPostfix := #tempPositionOfPostfix + 1;
       #tempPositionOfOperatorStack := #tempPositionOfOperatorStack - 1;
       #tempStackForOperators[#tempPositionOfOperatorStack] := #tempPrePostfix[#tempPositionOfPrePostfix];
       #tempPositionOfOperatorStack := #tempPositionOfOperatorStack + 1;
     ELSIF
       //kommende Öffnende Klammer ( immer in Zeichenspeicher speichern
       (#tempPrePostfix[#tempPositionOfPrePostfix] = #LGCODE_MTH_PRSR_OPEN_BRACKET)
     THEN
       #tempStackForOperators[#tempPositionOfOperatorStack] := #LGCODE_MTH_PRSR_OPEN_BRACKET;
       #tempPositionOfOperatorStack := #tempPositionOfOperatorStack + 1;
     ELSIF
       //letztes Zeichen eine öffnende Klammer (, dann kommendes Zeichen in Zeichenspeicher schreiben
       (#tempStackForOperators[#tempPositionOfOperatorStack - 1] = #LGCODE_MTH_PRSR_OPEN_BRACKET)
       AND
       ((#tempPrePostfix[#tempPositionOfPrePostfix] = #LGCODE_MTH_PRSR_LOGICAL_GREATER) OR
       (#tempPrePostfix[#tempPositionOfPrePostfix] = #LGCODE_MTH_PRSR_LOGICAL_LESS) OR
       (#tempPrePostfix[#tempPositionOfPrePostfix] = #LGCODE_MTH_PRSR_LOGICAL_GREATER_EQUAL) OR
       (#tempPrePostfix[#tempPositionOfPrePostfix] = #LGCODE_MTH_PRSR_LOGICAL_LESS_EQUAL) OR
       (#tempPrePostfix[#tempPositionOfPrePostfix] = #LGCODE_MTH_PRSR_LOGICAL_EQUAL) OR
       (#tempPrePostfix[#tempPositionOfPrePostfix] = #LGCODE_MTH_PRSR_LOGICAL_AND) OR
       (#tempPrePostfix[#tempPositionOfPrePostfix] = #LGCODE_MTH_PRSR_LOGICAL_OR) OR
       (#tempPrePostfix[#tempPositionOfPrePostfix] = #LGCODE_MTH_PRSR_PLUS) OR
       (#tempPrePostfix[#tempPositionOfPrePostfix] = #LGCODE_MTH_PRSR_MINUS) OR
       (#tempPrePostfix[#tempPositionOfPrePostfix] = #LGCODE_MTH_PRSR_TIMES) OR
       (#tempPrePostfix[#tempPositionOfPrePostfix] = #LGCODE_MTH_PRSR_DIVIDE))
     THEN
       #tempStackForOperators[#tempPositionOfOperatorStack] := #tempPrePostfix[#tempPositionOfPrePostfix];
       #tempPositionOfOperatorStack := #tempPositionOfOperatorStack + 1;
     ELSIF
       //nächstes Zeichen ist eine schließende Klammer
       //alle Zeichen aus Zeichenspeicher bis zur öffnenden Klammer in Postfix-Notation schreiben
       (#tempPrePostfix[#tempPositionOfPrePostfix] = #LGCODE_MTH_PRSR_CLOSE_BRACKET)
     THEN
       WHILE (#tempStackForOperators[#tempPositionOfOperatorStack - 1] <> #LGCODE_MTH_PRSR_OPEN_BRACKET) DO
         #tempPostfixNotation[#tempPositionOfPostfix] := #tempStackForOperators[#tempPositionOfOperatorStack - 1];
         #tempStackForOperators[#tempPositionOfOperatorStack - 1] := 0;
         #tempPositionOfOperatorStack := #tempPositionOfOperatorStack - 1;
         #tempPositionOfPostfix := #tempPositionOfPostfix + 1;
         //Falls eine negative mathematische Funktion kommt
         IF (#tempPositionOfNegFunctions[#tempNumberOfNegFunctions - 1] = #tempPositionOfOperatorStack) THEN
           #tempPositionOfNegTerm[#tempNumberOfNegTerm] := #tempPositionOfPostfix;
           #tempPositionOfPostfix := #tempPositionOfPostfix + 1;
           #tempNumberOfNegTerm := #tempNumberOfNegTerm + 1;
           #tempNumberOfNegFunctions := #tempNumberOfNegFunctions - 1;
         END_IF;
       END_WHILE;
       #tempPositionOfOperatorStack := #tempPositionOfOperatorStack - 1;
       #tempStackForOperators[#tempPositionOfOperatorStack] := 0;    //öffnende Klammer löschen
       //negative Klammerausdrücke
       IF (#tempPositionOfNegBrackets[#tempNumberOfNegBrackets - 1] = #tempPositionOfOperatorStack) THEN
         #tempPositionOfNegTerm[#tempNumberOfNegTerm] := #tempPositionOfPostfix;
         #tempPositionOfPostfix := #tempPositionOfPostfix + 1;
         #tempNumberOfNegTerm := #tempNumberOfNegTerm + 1;
         #tempNumberOfNegBrackets := #tempNumberOfNegBrackets - 1;
       END_IF;
     ELSIF    //sqr Quadrat
       (#tempPrePostfix[#tempPositionOfPrePostfix] = #LGCODE_MTH_PRSR_CHAR_S) AND
       (#tempPrePostfix[#tempPositionOfPrePostfix + 1] = #LGCODE_MTH_PRSR_CHAR_Q) AND
       (#tempPrePostfix[#tempPositionOfPrePostfix + 2] = #LGCODE_MTH_PRSR_CHAR_R) AND
       (#tempPrePostfix[#tempPositionOfPrePostfix + 3] <> #LGCODE_MTH_PRSR_CHAR_T)
     THEN
       #tempStackForOperators[#tempPositionOfOperatorStack] := #LGCODE_MTH_PRSR_SQUARE;
       #tempPositionOfOperatorStack := #tempPositionOfOperatorStack + 1;
       #tempPositionOfPrePostfix := #tempPositionOfPrePostfix + 2;
     ELSIF    //sqrt Quadratwurzel
       (#tempPrePostfix[#tempPositionOfPrePostfix] = #LGCODE_MTH_PRSR_CHAR_S) AND
       (#tempPrePostfix[#tempPositionOfPrePostfix + 1] = #LGCODE_MTH_PRSR_CHAR_Q) AND
       (#tempPrePostfix[#tempPositionOfPrePostfix + 2] = #LGCODE_MTH_PRSR_CHAR_R) AND
       (#tempPrePostfix[#tempPositionOfPrePostfix + 3] = #LGCODE_MTH_PRSR_CHAR_T)
     THEN
       #tempStackForOperators[#tempPositionOfOperatorStack] := #LGCODE_MTH_PRSR_SQUAREROOT;
       #tempPositionOfOperatorStack := #tempPositionOfOperatorStack + 1;
       #tempPositionOfPrePostfix := #tempPositionOfPrePostfix + 3;
     ELSIF    //sin Sinus
       (#tempPrePostfix[#tempPositionOfPrePostfix] = #LGCODE_MTH_PRSR_CHAR_S) AND
       (#tempPrePostfix[#tempPositionOfPrePostfix + 1] = #LGCODE_MTH_PRSR_CHAR_I) AND
       (#tempPrePostfix[#tempPositionOfPrePostfix + 2] = #LGCODE_MTH_PRSR_CHAR_N)
     THEN
       #tempStackForOperators[#tempPositionOfOperatorStack] := #LGCODE_MTH_PRSR_SINUS;
       #tempPositionOfOperatorStack := #tempPositionOfOperatorStack + 1;
       #tempPositionOfPrePostfix := #tempPositionOfPrePostfix + 2;
     ELSIF    //cos Cosinus
       (#tempPrePostfix[#tempPositionOfPrePostfix] = #LGCODE_MTH_PRSR_CHAR_C) AND
       (#tempPrePostfix[#tempPositionOfPrePostfix + 1] = #LGCODE_MTH_PRSR_CHAR_O) AND
       (#tempPrePostfix[#tempPositionOfPrePostfix + 2] = #LGCODE_MTH_PRSR_CHAR_S)
     THEN
       #tempStackForOperators[#tempPositionOfOperatorStack] := #LGCODE_MTH_PRSR_COSINUS;
       #tempPositionOfOperatorStack := #tempPositionOfOperatorStack + 1;
       #tempPositionOfPrePostfix := #tempPositionOfPrePostfix + 2;
     ELSIF
       //letztes Zeichen im Stack ist eine mathematische Funktion und Nächstes ein Rechen-Operator
       //Funktion wird auch bei logischen Operatoren (außer bei NOT) ausgelsen, oben realisiert
       ((#tempStackForOperators[#tempPositionOfOperatorStack - 1] = #LGCODE_MTH_PRSR_COSINUS) OR
       (#tempStackForOperators[#tempPositionOfOperatorStack - 1] = #LGCODE_MTH_PRSR_SINUS) OR
       (#tempStackForOperators[#tempPositionOfOperatorStack - 1] = #LGCODE_MTH_PRSR_SQUARE) OR
       (#tempStackForOperators[#tempPositionOfOperatorStack - 1] = #LGCODE_MTH_PRSR_SQUAREROOT)) AND
       ((#tempPrePostfix[#tempPositionOfPrePostfix] = #LGCODE_MTH_PRSR_TIMES) OR
       (#tempPrePostfix[#tempPositionOfPrePostfix] = #LGCODE_MTH_PRSR_MINUS) OR
       (#tempPrePostfix[#tempPositionOfPrePostfix] = #LGCODE_MTH_PRSR_PLUS) OR
       (#tempPrePostfix[#tempPositionOfPrePostfix] = #LGCODE_MTH_PRSR_DIVIDE))
     THEN
       #tempPostfixNotation[#tempPositionOfPostfix] := #tempStackForOperators[#tempPositionOfOperatorStack - 1];
       #tempPositionOfPostfix := #tempPositionOfPostfix + 1;
       #tempPositionOfOperatorStack := #tempPositionOfOperatorStack - 1;
       //Falls die mathematische Funktion negative ist
       IF (#tempPositionOfNegFunctions[#tempNumberOfNegFunctions - 1] = #tempPositionOfOperatorStack) THEN
         #tempPositionOfNegTerm[#tempNumberOfNegTerm] := #tempPositionOfPostfix;
         #tempPositionOfPostfix := #tempPositionOfPostfix + 1;
         #tempNumberOfNegTerm := #tempNumberOfNegTerm + 1;
         #tempNumberOfNegFunctions := #tempNumberOfNegFunctions - 1;
       END_IF;
       #tempPositionOfPrePostfix := #tempPositionOfPrePostfix - 1;
     ELSE
       ;
     END_IF;
     //Wenn PrePostfix-Array komplett eingelesen, Zeichenspeicher vollständig leeren
     IF (#tempPositionOfPrePostfix = #tempMaxPositionOfPrePostfix) THEN
       WHILE (#tempPositionOfOperatorStack > 1) DO
         #tempPostfixNotation[#tempPositionOfPostfix] := #tempStackForOperators[#tempPositionOfOperatorStack - 1];
         #tempStackForOperators[#tempPositionOfOperatorStack - 1] := 0;
         #tempPositionOfOperatorStack := #tempPositionOfOperatorStack - 1;
         #tempPositionOfPostfix := #tempPositionOfPostfix + 1;
         //Falls die mathematische Funktion negative ist
         IF (#tempPositionOfNegFunctions[#tempNumberOfNegFunctions - 1] = #tempPositionOfOperatorStack) THEN
           #tempPositionOfNegTerm[#tempNumberOfNegTerm] := #tempPositionOfPostfix;
           #tempPositionOfPostfix := #tempPositionOfPostfix + 1;
           #tempNumberOfNegTerm := #tempNumberOfNegTerm + 1;
           #tempNumberOfNegFunctions := #tempNumberOfNegFunctions - 1;
         END_IF;
       END_WHILE;
     END_IF;
     #tempPositionOfPrePostfix := #tempPositionOfPrePostfix + 1;
     #tempMaxOfPostfixPosition := #tempPositionOfPostfix;
   END_WHILE;
   #tempPositionOfPostfix := 1;
   #tempNumberOfMultiDigitNo := 1;
   #tempNumberOfNegTerm := 1;

   //Auswertung
   WHILE (#tempPositionOfPostfix <= #tempMaxOfPostfixPosition) DO
     IF (#tempPositionOfPostfix = #tempPositionOfNegTerm[#tempNumberOfNegTerm]) THEN
       //Vorzeichen des Ergebnisses des Klammerausdruckes negieren
       #tempStackOfIntermediateResults[#tempPositionOfIntermediateResult - 1] :=
       #tempStackOfIntermediateResults[#tempPositionOfIntermediateResult - 1] * (-1);
       #tempNumberOfNegTerm := #tempNumberOfNegTerm + 1;
       //Auswertung Zahlen Zeichen usw.
     ELSIF
       //um mehrstellige Zahlen nicht mit den ASCII Codierungen für Operatoren und Funktionen zu verwechseln
       (#tempPositionOfPostfix = #tempPositionMultiDigitNumbers[#tempNumberOfMultiDigitNo])
     THEN
       #tempStackOfIntermediateResults[#tempPositionOfIntermediateResult] := #tempPostfixNotation[#tempPositionOfPostfix];
       #tempPositionOfIntermediateResult := #tempPositionOfIntermediateResult + 1;
       #tempNumberOfMultiDigitNo := #tempNumberOfMultiDigitNo + 1;
     ELSIF
       //Falls Kommazahlen, negative Zahlen kommen, Abfrage kommendes Zeichen ungleich + - * /
       (#tempPostfixNotation[#tempPositionOfPostfix] <> #LGCODE_MTH_PRSR_LOGICAL_GREATER) AND
       (#tempPostfixNotation[#tempPositionOfPostfix] <> #LGCODE_MTH_PRSR_LOGICAL_LESS) AND
       (#tempPostfixNotation[#tempPositionOfPostfix] <> #LGCODE_MTH_PRSR_LOGICAL_GREATER_EQUAL) AND
       (#tempPostfixNotation[#tempPositionOfPostfix] <> #LGCODE_MTH_PRSR_LOGICAL_LESS_EQUAL) AND
       (#tempPostfixNotation[#tempPositionOfPostfix] <> #LGCODE_MTH_PRSR_LOGICAL_AND) AND
       (#tempPostfixNotation[#tempPositionOfPostfix] <> #LGCODE_MTH_PRSR_LOGICAL_OR) AND
       (#tempPostfixNotation[#tempPositionOfPostfix] <> #LGCODE_MTH_PRSR_LOGICAL_NOT) AND
       (#tempPostfixNotation[#tempPositionOfPostfix] <> #LGCODE_MTH_PRSR_LOGICAL_NOT_EQUAL) AND
       (#tempPostfixNotation[#tempPositionOfPostfix] <> #LGCODE_MTH_PRSR_LOGICAL_EQUAL) AND
       (#tempPostfixNotation[#tempPositionOfPostfix] <> #LGCODE_MTH_PRSR_MINUS) AND
       (#tempPostfixNotation[#tempPositionOfPostfix] <> #LGCODE_MTH_PRSR_PLUS) AND
       (#tempPostfixNotation[#tempPositionOfPostfix] <> #LGCODE_MTH_PRSR_TIMES) AND
       (#tempPostfixNotation[#tempPositionOfPostfix] <> #LGCODE_MTH_PRSR_DIVIDE) AND
       (#tempPostfixNotation[#tempPositionOfPostfix] <> #LGCODE_MTH_PRSR_SQUARE) AND
       (#tempPostfixNotation[#tempPositionOfPostfix] <> #LGCODE_MTH_PRSR_SQUAREROOT) AND
       (#tempPostfixNotation[#tempPositionOfPostfix] <> #LGCODE_MTH_PRSR_SINUS) AND
       (#tempPostfixNotation[#tempPositionOfPostfix] <> #LGCODE_MTH_PRSR_COSINUS) AND
       (#tempPostfixNotation[#tempPositionOfPostfix] <> #LGCODE_MTH_PRSR_TO_THE_POWER_OF)
     THEN
       #tempStackOfIntermediateResults[#tempPositionOfIntermediateResult] :=
       #tempPostfixNotation[#tempPositionOfPostfix];
       #tempPositionOfIntermediateResult := #tempPositionOfIntermediateResult + 1;

       //Auswertung ob +, -, * oder / und eigentliche Berechnung des mathematischen Ausdrucks
     ELSIF (#tempPostfixNotation[#tempPositionOfPostfix] = #LGCODE_MTH_PRSR_PLUS) THEN
       #tempStackOfIntermediateResults[#tempPositionOfIntermediateResult - 2] :=
       #tempStackOfIntermediateResults[#tempPositionOfIntermediateResult - 2] +
       #tempStackOfIntermediateResults[#tempPositionOfIntermediateResult - 1];
       #tempPositionOfIntermediateResult := #tempPositionOfIntermediateResult - 1;
     ELSIF (#tempPostfixNotation[#tempPositionOfPostfix] = #LGCODE_MTH_PRSR_MINUS) THEN
       #tempStackOfIntermediateResults[#tempPositionOfIntermediateResult - 2] :=
       #tempStackOfIntermediateResults[#tempPositionOfIntermediateResult - 2] -
       #tempStackOfIntermediateResults[#tempPositionOfIntermediateResult - 1];
       #tempPositionOfIntermediateResult := #tempPositionOfIntermediateResult - 1;
     ELSIF (#tempPostfixNotation[#tempPositionOfPostfix] = #LGCODE_MTH_PRSR_TIMES) THEN
       #tempStackOfIntermediateResults[#tempPositionOfIntermediateResult - 2] :=
       #tempStackOfIntermediateResults[#tempPositionOfIntermediateResult - 2] *
       #tempStackOfIntermediateResults[#tempPositionOfIntermediateResult - 1];
       #tempPositionOfIntermediateResult := #tempPositionOfIntermediateResult - 1;
     ELSIF (#tempPostfixNotation[#tempPositionOfPostfix] = #LGCODE_MTH_PRSR_DIVIDE) THEN

       // Prüfen auf Division durch Null
       IF (#tempStackOfIntermediateResults[#tempPositionOfIntermediateResult - 1] <> 0.0) THEN
         #tempStackOfIntermediateResults[#tempPositionOfIntermediateResult - 2] :=
         #tempStackOfIntermediateResults[#tempPositionOfIntermediateResult - 2] /
         #tempStackOfIntermediateResults[#tempPositionOfIntermediateResult - 1];
       ELSE
         #LKinLang_CalcMathAndBool.errorID := #LGCODE_MTH_PRSR_ERR_ID_DIVISION_BY_ZERO;
         #LKinLang_CalcMathAndBool.finalResult := 0;

         RETURN;
       END_IF;

       #tempPositionOfIntermediateResult := #tempPositionOfIntermediateResult - 1;
       //Auswertung sqr
     ELSIF (#tempPostfixNotation[#tempPositionOfPostfix] = #LGCODE_MTH_PRSR_SQUARE) THEN
       #tempStackOfIntermediateResults[#tempPositionOfIntermediateResult - 1] :=
       #tempStackOfIntermediateResults[#tempPositionOfIntermediateResult - 1] ** 2;
       //Auswertung sqrt
     ELSIF (#tempPostfixNotation[#tempPositionOfPostfix] = #LGCODE_MTH_PRSR_SQUAREROOT) THEN

       // Prüfen auf negative Wurzel
       IF (#tempStackOfIntermediateResults[#tempPositionOfIntermediateResult - 1] < 0.0) THEN
         #LKinLang_CalcMathAndBool.errorID := #LGCODE_MTH_PRSR_ERR_ID_NEAGTIVE_SQUARE_ROOT_ARGUMENT;
         #LKinLang_CalcMathAndBool.finalResult := 0;

         RETURN;
       ELSE
         #tempStackOfIntermediateResults[#tempPositionOfIntermediateResult - 1] :=
         SQRT(IN := #tempStackOfIntermediateResults[#tempPositionOfIntermediateResult - 1]);
       END_IF;

       //Auswertung sin
     ELSIF (#tempPostfixNotation[#tempPositionOfPostfix] = #LGCODE_MTH_PRSR_SINUS) THEN
       #tempStackOfIntermediateResults[#tempPositionOfIntermediateResult - 1] :=
       SIN(IN := #tempStackOfIntermediateResults[#tempPositionOfIntermediateResult - 1] * #LGCODE_MTH_PRSR_PI / 180);
       //Auswertung cos
     ELSIF (#tempPostfixNotation[#tempPositionOfPostfix] = #LGCODE_MTH_PRSR_COSINUS) THEN
       #tempStackOfIntermediateResults[#tempPositionOfIntermediateResult - 1] :=
       COS(IN := #tempStackOfIntermediateResults[#tempPositionOfIntermediateResult - 1] * #LGCODE_MTH_PRSR_PI / 180);
       //Auswertung Exponential-Rechnung
     ELSIF (#tempPostfixNotation[#tempPositionOfPostfix] = #LGCODE_MTH_PRSR_TO_THE_POWER_OF) THEN
       //Prüfen auf Einhaltung der SIMOTION Regeln für Exponential-Rechnung
       //1.Operand = 0, 2.Operand < 0
       IF (#tempStackOfIntermediateResults[#tempPositionOfIntermediateResult - 2] = 0.0) AND
         (#tempStackOfIntermediateResults[#tempPositionOfIntermediateResult - 1] < 0.0)
       THEN
         #LKinLang_CalcMathAndBool.errorID := #LGCODE_MTH_PRSR_ERR_ID_BASIS_ZERO_EXPONENT_NEGATIVE;
         #LKinLang_CalcMathAndBool.finalResult := 0;
         RETURN;
       ELSIF
         //Prüfen auf Einhaltung der SIMOTION Regeln für Exponential-Rechnung
         //1.Operand = 0, 2.Operand darf keine Dezimalzahl sein
         (#tempStackOfIntermediateResults[#tempPositionOfIntermediateResult - 2] < 0.0) AND
         ((#tempPositionOfPostfix - 1) = #tempPositionDecimalNumbers[#tempNumberOfDecimalNo])
       THEN
         #tempNumberOfDecimalNo := #tempNumberOfDecimalNo + 1;
         #LKinLang_CalcMathAndBool.errorID := #LGCODE_MTH_PRSR_ERR_ID_BASIS_NEGATIVE_EXPONENT_REAL;
         #LKinLang_CalcMathAndBool.finalResult := 0;
         RETURN;
       ELSE
         #tempStackOfIntermediateResults[#tempPositionOfIntermediateResult - 2] :=
         #tempStackOfIntermediateResults[#tempPositionOfIntermediateResult - 2] **
         #tempStackOfIntermediateResults[#tempPositionOfIntermediateResult - 1];
         #tempPositionOfIntermediateResult := #tempPositionOfIntermediateResult - 1;
       END_IF;
     ELSIF (#tempPostfixNotation[#tempPositionOfPostfix] = #LGCODE_MTH_PRSR_LOGICAL_GREATER) THEN
       IF
         #tempStackOfIntermediateResults[#tempPositionOfIntermediateResult - 2] >
         #tempStackOfIntermediateResults[#tempPositionOfIntermediateResult - 1]
       THEN
         #tempStackOfIntermediateResults[#tempPositionOfIntermediateResult - 2] := 1;
       ELSE
         #tempStackOfIntermediateResults[#tempPositionOfIntermediateResult - 2] := 0;
       END_IF;
       #tempPositionOfIntermediateResult := #tempPositionOfIntermediateResult - 1;

     ELSIF (#tempPostfixNotation[#tempPositionOfPostfix] = #LGCODE_MTH_PRSR_LOGICAL_LESS) THEN
       IF
         #tempStackOfIntermediateResults[#tempPositionOfIntermediateResult - 2] <
         #tempStackOfIntermediateResults[#tempPositionOfIntermediateResult - 1]
       THEN
         #tempStackOfIntermediateResults[#tempPositionOfIntermediateResult - 2] := 1;
       ELSE
         #tempStackOfIntermediateResults[#tempPositionOfIntermediateResult - 2] := 0;
       END_IF;
       #tempPositionOfIntermediateResult := #tempPositionOfIntermediateResult - 1;

     ELSIF (#tempPostfixNotation[#tempPositionOfPostfix] = #LGCODE_MTH_PRSR_LOGICAL_GREATER_EQUAL) THEN
       IF
         #tempStackOfIntermediateResults[#tempPositionOfIntermediateResult - 2] >=
         #tempStackOfIntermediateResults[#tempPositionOfIntermediateResult - 1]
       THEN
         #tempStackOfIntermediateResults[#tempPositionOfIntermediateResult - 2] := 1;
       ELSE
         #tempStackOfIntermediateResults[#tempPositionOfIntermediateResult - 2] := 0;
       END_IF;
       #tempPositionOfIntermediateResult := #tempPositionOfIntermediateResult - 1;

     ELSIF (#tempPostfixNotation[#tempPositionOfPostfix] = #LGCODE_MTH_PRSR_LOGICAL_LESS_EQUAL) THEN
       IF
         #tempStackOfIntermediateResults[#tempPositionOfIntermediateResult - 2] <=
         #tempStackOfIntermediateResults[#tempPositionOfIntermediateResult - 1]
       THEN
         #tempStackOfIntermediateResults[#tempPositionOfIntermediateResult - 2] := 1;
       ELSE
         #tempStackOfIntermediateResults[#tempPositionOfIntermediateResult - 2] := 0;
       END_IF;
       #tempPositionOfIntermediateResult := #tempPositionOfIntermediateResult - 1;